REGION Network 5: Procedure Selected
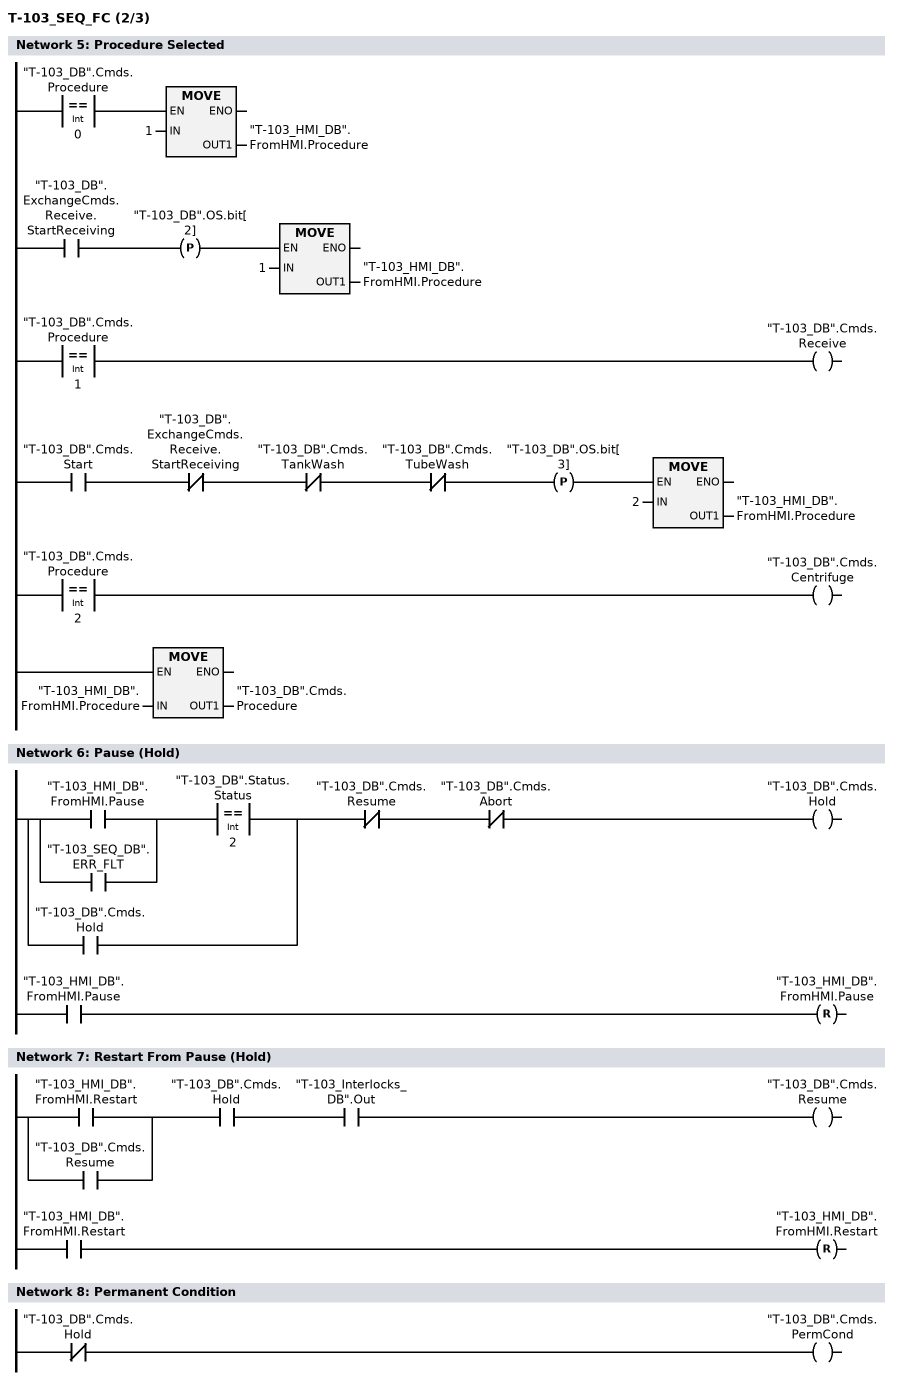
   RUNG wire#powerrail
      { S7_Templates := "SrcType := Int" } EQ_Contact(in1 := "T-103_DB".Cmds.Procedure, in2 := 0)
      Move(in := 1, out1 => "T-103_HMI_DB".FromHMI.Procedure)
   END_RUNG
   RUNG wire#powerrail
      Contact( "T-103_DB".ExchangeCmds.Receive.StartReceiving )
      P_Trig( "T-103_DB".OS.bit[2] )
      Move(in := 1, out1 => "T-103_HMI_DB".FromHMI.Procedure)
   END_RUNG
   RUNG wire#powerrail
      { S7_Templates := "SrcType := Int" } EQ_Contact(in1 := "T-103_DB".Cmds.Procedure, in2 := 1)
      Coil( "T-103_DB".Cmds.Receive )
   END_RUNG
   RUNG wire#powerrail
      Contact( "T-103_DB".Cmds.Start )
      I_Contact( "T-103_DB".ExchangeCmds.Receive.StartReceiving )
      I_Contact( "T-103_DB".Cmds.TankWash )
      I_Contact( "T-103_DB".Cmds.TubeWash )
      P_Trig( "T-103_DB".OS.bit[3] )
      Move(in := 2, out1 => "T-103_HMI_DB".FromHMI.Procedure)
   END_RUNG
   RUNG wire#powerrail
      { S7_Templates := "SrcType := Int" } EQ_Contact(in1 := "T-103_DB".Cmds.Procedure, in2 := 2)
      Coil( "T-103_DB".Cmds.Centrifuge )
   END_RUNG
   RUNG wire#powerrail
      Move(in := "T-103_HMI_DB".FromHMI.Procedure, out1 => "T-103_DB".Cmds.Procedure)
   END_RUNG
   // the same network as SCL:
   IF "T-103_DB".Cmds.Procedure = 0 THEN "T-103_HMI_DB".FromHMI.Procedure := 1; END_IF;
   #_w1 := "T-103_DB".ExchangeCmds.Receive.StartReceiving AND NOT "T-103_DB".OS.bit[2];   // rising edge
   "T-103_DB".OS.bit[2] := "T-103_DB".ExchangeCmds.Receive.StartReceiving;
   IF #_w1 THEN "T-103_HMI_DB".FromHMI.Procedure := 1; END_IF;
   "T-103_DB".Cmds.Receive := "T-103_DB".Cmds.Procedure = 1;
   #_w2 := "T-103_DB".Cmds.Start AND NOT "T-103_DB".ExchangeCmds.Receive.StartReceiving AND NOT "T-103_DB".Cmds.TankWash AND NOT "T-103_DB".Cmds.TubeWash;
   #_w3 := #_w2 AND NOT "T-103_DB".OS.bit[3];   // rising edge
   "T-103_DB".OS.bit[3] := #_w2;
   IF #_w3 THEN "T-103_HMI_DB".FromHMI.Procedure := 2; END_IF;
   "T-103_DB".Cmds.Centrifuge := "T-103_DB".Cmds.Procedure = 2;
   "T-103_DB".Cmds.Procedure := "T-103_HMI_DB".FromHMI.Procedure;
END_REGION

REGION Network 6: Pause (Hold)
   RUNG wire#powerrail
      Contact( "T-103_HMI_DB".FromHMI.Pause )
      wire#w1
      { S7_Templates := "SrcType := Int" } EQ_Contact(in1 := "T-103_DB".Status.Status, in2 := 2)
      wire#w2
      I_Contact( "T-103_DB".Cmds.Resume )
      I_Contact( "T-103_DB".Cmds.Abort )
      Coil( "T-103_DB".Cmds.Hold )
   END_RUNG
   RUNG wire#powerrail
      Contact( "T-103_SEQ_DB".ERR_FLT )
   END_RUNG wire#w1
   RUNG wire#powerrail
      Contact( "T-103_DB".Cmds.Hold )
   END_RUNG wire#w2
   RUNG wire#powerrail
      Contact( "T-103_HMI_DB".FromHMI.Pause )
      R_Coil( "T-103_HMI_DB".FromHMI.Pause )
   END_RUNG
   // the same network as SCL:
   "T-103_DB".Cmds.Hold := ((("T-103_HMI_DB".FromHMI.Pause OR "T-103_SEQ_DB".ERR_FLT) AND ("T-103_DB".Status.Status = 2)) OR "T-103_DB".Cmds.Hold) AND NOT "T-103_DB".Cmds.Resume AND NOT "T-103_DB".Cmds.Abort;
   IF "T-103_HMI_DB".FromHMI.Pause THEN "T-103_HMI_DB".FromHMI.Pause := FALSE; END_IF;
END_REGION

REGION Network 7: Restart From Pause (Hold)
   RUNG wire#powerrail
      Contact( "T-103_HMI_DB".FromHMI.Restart )
      wire#w1
      Contact( "T-103_DB".Cmds.Hold )
      Contact( "T-103_Interlocks_DB".Out )
      Coil( "T-103_DB".Cmds.Resume )
   END_RUNG
   RUNG wire#powerrail
      Contact( "T-103_DB".Cmds.Resume )
   END_RUNG wire#w1
   RUNG wire#powerrail
      Contact( "T-103_HMI_DB".FromHMI.Restart )
      R_Coil( "T-103_HMI_DB".FromHMI.Restart )
   END_RUNG
   // the same network as SCL:
   "T-103_DB".Cmds.Resume := ("T-103_HMI_DB".FromHMI.Restart OR "T-103_DB".Cmds.Resume) AND "T-103_DB".Cmds.Hold AND "T-103_Interlocks_DB".Out;
   IF "T-103_HMI_DB".FromHMI.Restart THEN "T-103_HMI_DB".FromHMI.Restart := FALSE; END_IF;
END_REGION

REGION Network 8: Permanent Condition
   RUNG wire#powerrail
      I_Contact( "T-103_DB".Cmds.Hold )
      Coil( "T-103_DB".Cmds.PermCond )
   END_RUNG
   // the same network as SCL:
   "T-103_DB".Cmds.PermCond := NOT "T-103_DB".Cmds.Hold;
END_REGION

REGION Network 9: Tank Wash
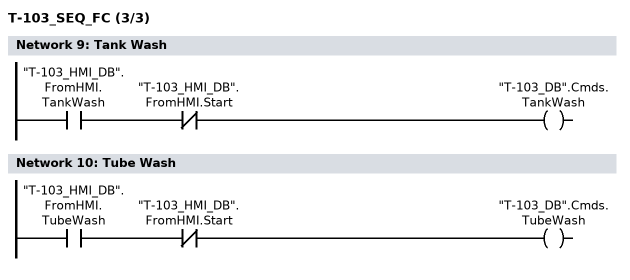
   RUNG wire#powerrail
      Contact( "T-103_HMI_DB".FromHMI.TankWash )
      I_Contact( "T-103_HMI_DB".FromHMI.Start )
      Coil( "T-103_DB".Cmds.TankWash )
   END_RUNG
   // the same network as SCL:
   "T-103_DB".Cmds.TankWash := "T-103_HMI_DB".FromHMI.TankWash AND NOT "T-103_HMI_DB".FromHMI.Start;
END_REGION

REGION Network 10: Tube Wash
   RUNG wire#powerrail
      Contact( "T-103_HMI_DB".FromHMI.TubeWash )
      I_Contact( "T-103_HMI_DB".FromHMI.Start )
      Coil( "T-103_DB".Cmds.TubeWash )
   END_RUNG
   // the same network as SCL:
   "T-103_DB".Cmds.TubeWash := "T-103_HMI_DB".FromHMI.TubeWash AND NOT "T-103_HMI_DB".FromHMI.Start;
END_REGION

REGION Network 11 (SCL): Sequence Status
   IF "T-103_SEQ_DB".S_NO= 1 THEN
       "T-103_DB".Status.Status := 1; //Idle
   ELSIF ("T-103_SEQ_DB".S_NO > 1 AND "T-103_SEQ_DB".S_NO < 150) AND NOT "T-103_SEQ_DB".ERR_FLT AND NOT "T-103_DB".Cmds.Hold THEN
       "T-103_DB".Status.Status := 2; //Running
   ELSIF "T-103_SEQ_DB".S_NO >= 151 AND "T-103_SEQ_DB".S_NO <= 160 AND NOT "T-103_SEQ_DB".ERR_FLT THEN
       "T-103_DB".Status.Status := 3; // Stopping
   ELSIF  "T-103_SEQ_DB".ERR_FLT AND  ("T-103_SEQ_DB".S_NO > 1 AND "T-103_SEQ_DB".S_NO < 150) THEN
       "T-103_DB".Status.Status := 4; // Held
   ELSIF  "T-103_SEQ_DB".ERR_FLT AND  ("T-103_SEQ_DB".S_NO > 1 AND "T-103_SEQ_DB".S_NO < 150) AND "T-103_Aux_DB"."Bool".TOff  THEN
       "T-103_DB".Status.Status := 5; // Holding
   ELSE
       "T-103_DB".Status.Status := 6; // Unknown
   END_IF;

   "T-103_DB".Status.Running := ("T-103_SEQ_DB".S_NO > 3 AND "T-103_SEQ_DB".S_NO <= 150);
   "T-103_DB".Status.Initializing := ("T-103_SEQ_DB".S_NO >= 141 AND "T-103_SEQ_DB".S_NO <= 150);

   //Enable/Disable HMI Start/Stop Button
   "T-103_HMI_DB".ToHMI.EnStopButton := ("T-103_DB".Status.Status > 1) OR "T-103_DB".Status.Step = 0; //Enable HMI Stop Button
   "T-103_HMI_DB".ToHMI.EnStartButton := "T-103_DB".Status.Status = 1; //Idle
   "T-103_HMI_DB".ToHMI.EnPauseButton := "T-103_DB".Status.Status = 2; //Enable Pause Button
   "T-103_HMI_DB".ToHMI.EnRestartButton :=  "T-103_DB".Status.Status = 4; //Enable Restart Button

   //****Interlock Activated
   "T-103_HMI_DB".ToHMI.InterlockActivated := "T-103_Interlocks_DB".Out;
END_REGION

REGION Network 12 (SCL): Sequence Step
   "T-103_DB".Status.Step := "T-103_SEQ_DB".S_NO;
END_REGION

REGION Network 13 (SCL): Sequence state (Procedure running)
   IF "T-103_SEQ_DB".S_NO = 3 OR "T-103_SEQ_DB".S_NO = 4 THEN
       "T-103_DB".Status.State := 1; //Ready
   ELSIF "T-103_SEQ_DB".S_NO >= 21 AND "T-103_SEQ_DB".S_NO <= 60 THEN
       "T-103_DB".Status.State := 2; //Mixing 
   ELSIF "T-103_SEQ_DB".S_NO >= 61 AND "T-103_SEQ_DB".S_NO <= 80 THEN
       "T-103_DB".Status.State := 3; //Pouring
   ELSIF "T-103_SEQ_DB".S_NO >= 141 AND "T-103_SEQ_DB".S_NO <= 150 THEN
       "T-103_DB".Status.State := 4; //Initializing
   ELSIF "T-103_SEQ_DB".S_NO >= 151 AND "T-103_SEQ_DB".S_NO <= 160 THEN
       "T-103_DB".Status.State := 5; //Aborting
   ELSE
       "T-103_DB".Status.State := 0;
   END_IF;
END_REGION

REGION Network 14: Sequence State
END_REGION
END_FUNCTION

// folder: State MACHINE/1)Tanks/Tank T-103 (Cooling Tank)/T-103 <---> Centrifuge

FUNCTION "T-103_Signals_FROM_Centrifuge" : Void   // FC69, LAD
{ S7_Optimized_Access := 'TRUE' }
VERSION : 0.1
BEGIN

REGION Network 1: Start Sequence
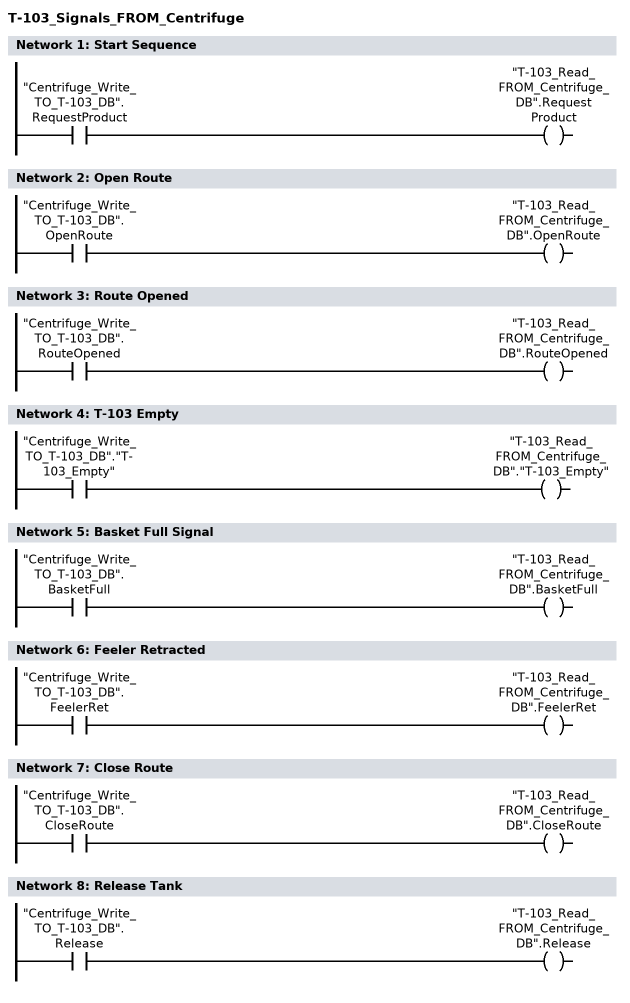
   RUNG wire#powerrail
      Contact( "Centrifuge_Write_TO_T-103_DB".RequestProduct )
      Coil( "T-103_Read_FROM_Centrifuge_DB".RequestProduct )
   END_RUNG
   // the same network as SCL:
   "T-103_Read_FROM_Centrifuge_DB".RequestProduct := "Centrifuge_Write_TO_T-103_DB".RequestProduct;
END_REGION

REGION Network 2: Open Route
   RUNG wire#powerrail
      Contact( "Centrifuge_Write_TO_T-103_DB".OpenRoute )
      Coil( "T-103_Read_FROM_Centrifuge_DB".OpenRoute )
   END_RUNG
   // the same network as SCL:
   "T-103_Read_FROM_Centrifuge_DB".OpenRoute := "Centrifuge_Write_TO_T-103_DB".OpenRoute;
END_REGION

REGION Network 3: Route Opened
   RUNG wire#powerrail
      Contact( "Centrifuge_Write_TO_T-103_DB".RouteOpened )
      Coil( "T-103_Read_FROM_Centrifuge_DB".RouteOpened )
   END_RUNG
   // the same network as SCL:
   "T-103_Read_FROM_Centrifuge_DB".RouteOpened := "Centrifuge_Write_TO_T-103_DB".RouteOpened;
END_REGION

REGION Network 4: T-103 Empty
   RUNG wire#powerrail
      Contact( "Centrifuge_Write_TO_T-103_DB"."T-103_Empty" )
      Coil( "T-103_Read_FROM_Centrifuge_DB"."T-103_Empty" )
   END_RUNG
   // the same network as SCL:
   "T-103_Read_FROM_Centrifuge_DB"."T-103_Empty" := "Centrifuge_Write_TO_T-103_DB"."T-103_Empty";
END_REGION

REGION Network 5: Basket Full Signal
   RUNG wire#powerrail
      Contact( "Centrifuge_Write_TO_T-103_DB".BasketFull )
      Coil( "T-103_Read_FROM_Centrifuge_DB".BasketFull )
   END_RUNG
   // the same network as SCL:
   "T-103_Read_FROM_Centrifuge_DB".BasketFull := "Centrifuge_Write_TO_T-103_DB".BasketFull;
END_REGION

REGION Network 6: Feeler Retracted
   RUNG wire#powerrail
      Contact( "Centrifuge_Write_TO_T-103_DB".FeelerRet )
      Coil( "T-103_Read_FROM_Centrifuge_DB".FeelerRet )
   END_RUNG
   // the same network as SCL:
   "T-103_Read_FROM_Centrifuge_DB".FeelerRet := "Centrifuge_Write_TO_T-103_DB".FeelerRet;
END_REGION

REGION Network 7: Close Route
   RUNG wire#powerrail
      Contact( "Centrifuge_Write_TO_T-103_DB".CloseRoute )
      Coil( "T-103_Read_FROM_Centrifuge_DB".CloseRoute )
   END_RUNG
   // the same network as SCL:
   "T-103_Read_FROM_Centrifuge_DB".CloseRoute := "Centrifuge_Write_TO_T-103_DB".CloseRoute;
END_REGION

REGION Network 8: Release Tank
   RUNG wire#powerrail
      Contact( "Centrifuge_Write_TO_T-103_DB".Release )
      Coil( "T-103_Read_FROM_Centrifuge_DB".Release )
   END_RUNG
   // the same network as SCL:
   "T-103_Read_FROM_Centrifuge_DB".Release := "Centrifuge_Write_TO_T-103_DB".Release;
END_REGION
END_FUNCTION

// folder: State MACHINE/1)Tanks/Tank T-103 (Cooling Tank)/T-103 <---> R-201

FUNCTION "T-103_Signals_FROM_R-201" : Void   // FC49, LAD
{ S7_Optimized_Access := 'TRUE' }
VERSION : 0.1
BEGIN

REGION Network 1: Start Sequence
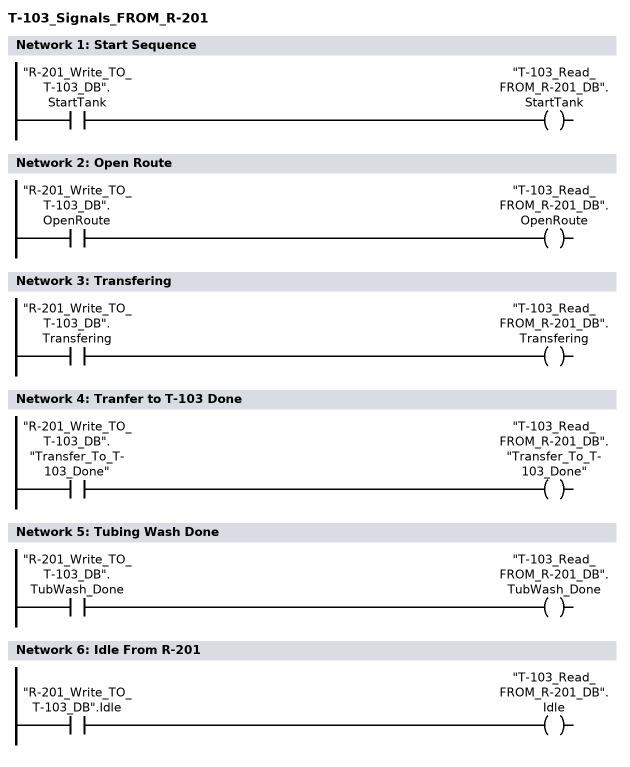
   RUNG wire#powerrail
      Contact( "R-201_Write_TO_T-103_DB".StartTank )
      Coil( "T-103_Read_FROM_R-201_DB".StartTank )
   END_RUNG
   // the same network as SCL:
   "T-103_Read_FROM_R-201_DB".StartTank := "R-201_Write_TO_T-103_DB".StartTank;
END_REGION

REGION Network 2: Open Route
   RUNG wire#powerrail
      Contact( "R-201_Write_TO_T-103_DB".OpenRoute )
      Coil( "T-103_Read_FROM_R-201_DB".OpenRoute )
   END_RUNG
   // the same network as SCL:
   "T-103_Read_FROM_R-201_DB".OpenRoute := "R-201_Write_TO_T-103_DB".OpenRoute;
END_REGION

REGION Network 3: Transfering
   RUNG wire#powerrail
      Contact( "R-201_Write_TO_T-103_DB".Transfering )
      Coil( "T-103_Read_FROM_R-201_DB".Transfering )
   END_RUNG
   // the same network as SCL:
   "T-103_Read_FROM_R-201_DB".Transfering := "R-201_Write_TO_T-103_DB".Transfering;
END_REGION

REGION Network 4: Tranfer to T-103 Done
   RUNG wire#powerrail
      Contact( "R-201_Write_TO_T-103_DB"."Transfer_To_T-103_Done" )
      Coil( "T-103_Read_FROM_R-201_DB"."Transfer_To_T-103_Done" )
   END_RUNG
   // the same network as SCL:
   "T-103_Read_FROM_R-201_DB"."Transfer_To_T-103_Done" := "R-201_Write_TO_T-103_DB"."Transfer_To_T-103_Done";
END_REGION

REGION Network 5: Tubing Wash Done
   RUNG wire#powerrail
      Contact( "R-201_Write_TO_T-103_DB".TubWash_Done )
      Coil( "T-103_Read_FROM_R-201_DB".TubWash_Done )
   END_RUNG
   // the same network as SCL:
   "T-103_Read_FROM_R-201_DB".TubWash_Done := "R-201_Write_TO_T-103_DB".TubWash_Done;
END_REGION

REGION Network 6: Idle From R-201
   RUNG wire#powerrail
      Contact( "R-201_Write_TO_T-103_DB".Idle )
      Coil( "T-103_Read_FROM_R-201_DB".Idle )
   END_RUNG
   // the same network as SCL:
   "T-103_Read_FROM_R-201_DB".Idle := "R-201_Write_TO_T-103_DB".Idle;
END_REGION
END_FUNCTION

// folder: State MACHINE/1)Tanks/Tank T-103 (Cooling Tank)/T-103 <--->R-202

FUNCTION "T-103_Signals_FROM_R-202" : Void   // FC63, LAD
{ S7_Optimized_Access := 'TRUE' }
VERSION : 0.1
BEGIN

REGION Network 1: Start Sequence
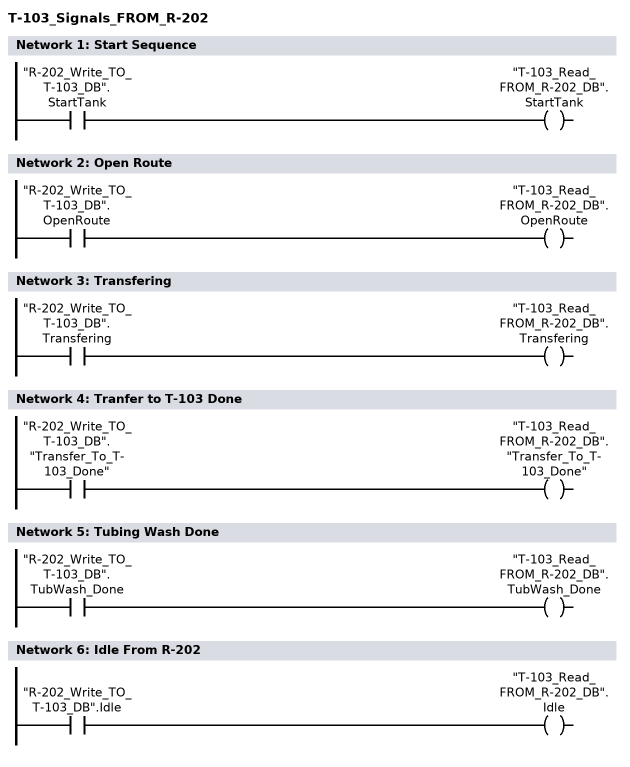
   RUNG wire#powerrail
      Contact( "R-202_Write_TO_T-103_DB".StartTank )
      Coil( "T-103_Read_FROM_R-202_DB".StartTank )
   END_RUNG
   // the same network as SCL:
   "T-103_Read_FROM_R-202_DB".StartTank := "R-202_Write_TO_T-103_DB".StartTank;
END_REGION

REGION Network 2: Open Route
   RUNG wire#powerrail
      Contact( "R-202_Write_TO_T-103_DB".OpenRoute )
      Coil( "T-103_Read_FROM_R-202_DB".OpenRoute )
   END_RUNG
   // the same network as SCL:
   "T-103_Read_FROM_R-202_DB".OpenRoute := "R-202_Write_TO_T-103_DB".OpenRoute;
END_REGION

REGION Network 3: Transfering
   RUNG wire#powerrail
      Contact( "R-202_Write_TO_T-103_DB".Transfering )
      Coil( "T-103_Read_FROM_R-202_DB".Transfering )
   END_RUNG
   // the same network as SCL:
   "T-103_Read_FROM_R-202_DB".Transfering := "R-202_Write_TO_T-103_DB".Transfering;
END_REGION

REGION Network 4: Tranfer to T-103 Done
   RUNG wire#powerrail
      Contact( "R-202_Write_TO_T-103_DB"."Transfer_To_T-103_Done" )
      Coil( "T-103_Read_FROM_R-202_DB"."Transfer_To_T-103_Done" )
   END_RUNG
   // the same network as SCL:
   "T-103_Read_FROM_R-202_DB"."Transfer_To_T-103_Done" := "R-202_Write_TO_T-103_DB"."Transfer_To_T-103_Done";
END_REGION

REGION Network 5: Tubing Wash Done
   RUNG wire#powerrail
      Contact( "R-202_Write_TO_T-103_DB".TubWash_Done )
      Coil( "T-103_Read_FROM_R-202_DB".TubWash_Done )
   END_RUNG
   // the same network as SCL:
   "T-103_Read_FROM_R-202_DB".TubWash_Done := "R-202_Write_TO_T-103_DB".TubWash_Done;
END_REGION

REGION Network 6: Idle From R-202
   RUNG wire#powerrail
      Contact( "R-202_Write_TO_T-103_DB".Idle )
      Coil( "T-103_Read_FROM_R-202_DB".Idle )
   END_RUNG
   // the same network as SCL:
   "T-103_Read_FROM_R-202_DB".Idle := "R-202_Write_TO_T-103_DB".Idle;
END_REGION
END_FUNCTION

// folder: State MACHINE/1)Tanks/Tank T-104 (Water System)

FUNCTION_BLOCK "T-104_SEQ"   // FB38, GRAPH_PLUS
{ S7_Optimized_Access := 'TRUE' }
VERSION : 0.1
   VAR_INPUT
      OFF_SQ : Bool := false;   // Turn sequence off
      INIT_SQ : Bool := false;   // Set sequence to initial state
      ACK_EF : Bool := false;   // Acknowledge all errors and faults
   END_VAR
   VAR_OUTPUT
      S_NO : Int := 0;   // Step number
      S_MORE : Bool := false;   // More steps are available and can be shown in S_NO
      S_ACTIVE : Bool := false;   // Step indicated in S_NO is active
      ERR_FLT : Bool := false;   // Interlock or supervision group error
      AUTO_ON : Bool := false;   // Automatic mode is active
   END_VAR
   VAR
      STATE : Int;   // Current Step in Sequence
      Tank : Struct   // Reactor Ctrl
         IDLE : Bool;
         INITIALIZATION : Bool;   // Sequence initialization
         START : Bool;
         DONE_REACTING : Bool;
         COMPLETE : Bool;   // Reactor Complete Read only
         PARA : Bool;   // PARA load Batch side button
         ABORTING : Bool;   // Sequence about
         WAIT : Bool;   // Wating for Permissive read only
      END_STRUCT;
      TEMP : Struct
         TANKS_BATCH : Real;
         "EMPTY_LV_0%" : Real;
         "MIN_LV_20%" : Real;
         "MAX_LV_80%" : Real;
         "BELOW_32%" : Real;
         "Greater_8%" : Real;
         "PRE-ADD" : Real;
         X_SOL_SIZE : Real;
         Y_SOL_SIZE : Real;
         OFFSEt : Struct
            MAX : Real;
            MIN : Real;
         END_STRUCT;
      END_STRUCT;
      HMI_INFO : Array[0..11] of UInt;
      IF_PAR : G7_IfParPlus_V6;
      RT_DATA : G7_RTDataPlus_V6;   // Internal data area
      Abort : G7_TransitionPlus_V6;   // Transition structure
      InitializeTk : G7_TransitionPlus_V6;   // Transition structure
      Block : G7_TransitionPlus_V6;   // Transition structure
      Rdy : G7_TransitionPlus_V6;   // Transition structure
      Feed : G7_TransitionPlus_V6;   // Transition structure
      ReqWater1 : G7_TransitionPlus_V6;   // Transition structure
      StopWater1 : G7_TransitionPlus_V6;   // Transition structure
      Stoped1 : G7_TransitionPlus_V6;   // Transition structure
      GoBack : G7_TransitionPlus_V6;   // Transition structure
      Init : G7_TransitionPlus_V6;   // Transition structure
      SAut : G7_TransitionPlus_V6;   // Transition structure
      SIn : G7_TransitionPlus_V6;   // Transition structure
      Initd : G7_TransitionPlus_V6;   // Transition structure
      Ab : G7_TransitionPlus_V6;   // Transition structure
      AbortOn : G7_TransitionPlus_V6;   // Transition structure
      DneAbort : G7_TransitionPlus_V6;   // Transition structure
      Idle : G7_StepPlus_V6;   // Step structure
      Ready : G7_StepPlus_V6;   // Step structure
      SelectSeq : G7_StepPlus_V6;   // Step structure
      FeedStarted : G7_StepPlus_V6;   // Step structure
      Feeding : G7_StepPlus_V6;   // Step structure
      StopTransfer : G7_StepPlus_V6;   // Step structure
      Done : G7_StepPlus_V6;   // Step structure
      Initialize : G7_StepPlus_V6;   // Step structure
      SetAuto : G7_StepPlus_V6;   // Step structure
      SetInitial : G7_StepPlus_V6;   // Step structure
      Initialized : G7_StepPlus_V6;   // Step structure
      AbortStarting : G7_StepPlus_V6;   // Step structure
      Aborting : G7_StepPlus_V6;   // Step structure
      Abort_Done : G7_StepPlus_V6;   // Step structure
      SINI : Array[0..4] of USInt;
      LSTT : Array[0..15] of USInt;
      ATAJ : Array[0..15] of USInt;
      ATAB : Array[0..15] of USInt;
      PSTT : Array[0..15] of USInt;
      NSTT : Array[0..15] of USInt;
      ASSJ : Array[0..13] of USInt;
      ASSB : Array[0..13] of USInt;
      PTTS : Array[0..13] of USInt;
      NTTS : Array[0..13] of USInt;
      SW_SQTS : Array[0..13] of USInt;
      SWITCH : Array[0..3] of USInt;
      TVX : Array[0..7] of USInt;
      TTX : Array[0..7] of USInt;
      TSX : Array[0..4] of USInt;
      S00X : Array[0..4] of USInt;
      SOFFX : Array[0..4] of USInt;
      SONX : Array[0..4] of USInt;
      SAX : Array[0..4] of USInt;
      SERRX : Array[0..14] of USInt;
      SMX : Array[0..14] of USInt;
      S0X : Array[0..14] of USInt;
      S1X : Array[0..14] of USInt;
      IL_ALARM_INST : Diag_Alarm;
      SUP_ALARM_INST : Diag_Alarm;
      STEP_TIME_ALARM_INST : Diag_Alarm;
      IEC_TIMER_INST : IEC_TIMER;
      TRANSACTION_FLAG : Bool := false;
   END_VAR
   VAR CONSTANT
      "Single R-201 T-101 seq done" : Int := 214;
      "Single R-201 T-102 seq done" : Int := 218;
   END_VAR
   // SINI[0] := 2;
   // LSTT[0] := 11;
   // NSTT[0] := 11;
   // PTTS[0] := 255;
   // TVX[0] := 16#1;
   // TTX[0] := 16#1;
   // TSX[0] := 16#1;
   // S00X[0] := 16#1;
   // SOFFX[0] := 16#1;
   // SONX[0] := 16#1;
   // SAX[0] := 16#1;
   // SERRX[0] := 16#1;
   // SMX[0] := 16#1;
   // S0X[0] := 16#1;
   // S1X[0] := 16#1;
   // LSTT[1] := 7;
   // LSTT[2] := 255;
   // LSTT[3] := 255;
   // LSTT[4] := 3;
   // LSTT[5] := 255;
   // LSTT[6] := 255;
   // LSTT[7] := 255;
   // LSTT[8] := 3;
   // LSTT[9] := 255;
   // LSTT[10] := 255;
   // LSTT[11] := 255;
   // LSTT[13] := 255;
   // ATAJ[1] := 1;
   // ATAJ[2] := 2;
   // ATAJ[3] := 3;
   // ATAJ[4] := 4;
   // ATAJ[5] := 5;
   // ATAJ[6] := 6;
   // ATAJ[7] := 7;
   // ATAJ[8] := 8;
   // ATAJ[9] := 9;
   // ATAJ[10] := 10;
   // ATAJ[11] := 11;
   // ATAJ[12] := 12;
   // ATAJ[13] := 13;
   // ATAB[1] := 2;
   // ATAB[13] := 13;
   // ATAB[3] := 3;
   // ATAB[4] := 4;
   // ATAB[5] := 5;
   // ATAB[6] := 6;
   // ATAB[7] := 7;
   // ATAB[8] := 8;
   // ATAB[9] := 9;
   // ATAB[10] := 10;
   // ATAB[11] := 11;
   // ATAB[12] := 12;
   // PSTT[3] := 1;
   // PSTT[4] := 2;
   // PSTT[5] := 3;
   // PSTT[6] := 4;
   // PSTT[7] := 5;
   // PSTT[8] := 6;
   // PSTT[9] := 7;
   // PSTT[10] := 8;
   // PSTT[11] := 9;
   // PSTT[12] := 10;
   // NSTT[1] := 7;
   // NSTT[2] := 1;
   // NSTT[3] := 2;
   // NSTT[4] := 3;
   // NSTT[5] := 4;
   // NSTT[6] := 5;
   // NSTT[7] := 6;
   // NSTT[8] := 3;
   // NSTT[9] := 8;
   // NSTT[10] := 9;
   // NSTT[11] := 10;
   // NSTT[13] := 12;
   // ASSJ[1] := 1;
   // ASSJ[2] := 2;
   // ASSJ[3] := 3;
   // ASSJ[4] := 4;
   // ASSJ[5] := 5;
   // ASSJ[6] := 6;
   // ASSJ[7] := 7;
   // ASSJ[8] := 8;
   // ASSJ[9] := 9;
   // ASSJ[10] := 10;
   // ASSJ[11] := 11;
   // ASSB[1] := 1;
   // ASSB[2] := 2;
   // ASSB[3] := 3;
   // ASSB[4] := 4;
   // ASSB[5] := 5;
   // ASSB[6] := 6;
   // ASSB[7] := 7;
   // ASSB[8] := 8;
   // ASSB[9] := 9;
   // ASSB[10] := 10;
   // ASSB[11] := 11;
   // PTTS[4] := 5;
   // PTTS[3] := 255;
   // PTTS[5] := 6;
   // PTTS[6] := 7;
   // PTTS[7] := 255;
   // PTTS[8] := 9;
   // PTTS[9] := 10;
   // PTTS[11] := 255;
   // SW_SQTS[4] := 2;
   // NTTS[2] := 4;
   // NTTS[3] := 5;
   // NTTS[4] := 6;
   // NTTS[5] := 7;
   // NTTS[6] := 8;
   // NTTS[7] := 9;
   // NTTS[8] := 10;
   // NTTS[9] := 11;
   // NTTS[10] := 12;
   // NTTS[11] := 13;
   // SW_SQTS[5] := 2;
   // SW_SQTS[8] := 3;
   // SW_SQTS[9] := 3;
   // SW_SQTS[11] := 4;
   // SWITCH[0] := 156;
   // SWITCH[2] := 251;
   // PSTT[13] := 11;
   // PTTS[1] := 2;
   // NTTS[1] := 3;
   // SW_SQTS[1] := 1;
   // PTTS[10] := 11;
   // ATAB[0] := 1;
   // SINI[4] := 255;
   // SINI[3] := 255;
   // PTTS[2] := 3;
   // SW_SQTS[7] := 3;
   // SW_SQTS[6] := 2;
   // SWITCH[1] := 239;
   // SINI[2] := 255;
   // SW_SQTS[3] := 2;
   // SW_SQTS[2] := 1;
   // SW_SQTS[10] := 3;
   // LSTT[12] := 1;
   // LSTT[14] := 255;
   // ATAJ[14] := 14;
   // ATAJ[15] := 15;
   // ATAB[14] := 14;
   // ATAB[15] := 15;
   // PSTT[14] := 12;
   // PSTT[15] := 13;
   // NSTT[12] := 1;
   // NSTT[14] := 13;
   // ASSJ[12] := 12;
   // ASSJ[13] := 13;
   // ASSB[12] := 12;
   // ASSB[13] := 13;
   // PTTS[12] := 13;
   // PTTS[13] := 14;
   // NTTS[12] := 14;
   // NTTS[13] := 15;
   // SW_SQTS[12] := 4;
   // SW_SQTS[13] := 4;
BEGIN
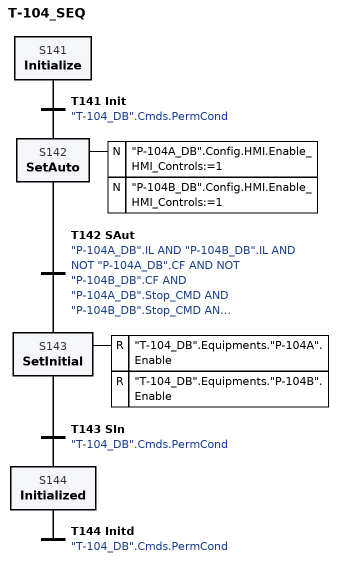
   // permanent pre-instructions
   NETWORK 1
      "T-104_SEQ_FC"();
      "T-104_Signals_FROM_R-201"();
      "T-104_Signals_FROM_R-202"();
      "T-104_Signals_FROM_T-101"();
      "T-104_Signals_FROM_T-102"();
      "T-104_Signals_FROM_Centrifuge"();
      "T-104_SignalsInExchange"();

   // sequencer 1
   STEP SetAuto:   // S142, max time T#10S, warning time T#7S
      // PMP OFF
              N    "P-104A_DB".Config.HMI.Enable_HMI_Controls:=1
              N    "P-104B_DB".Config.HMI.Enable_HMI_Controls:=1
   END_STEP
   TRANSITION SAut FROM SetAuto TO SetInitial   // T142: OFF: P-101A/B
      := "P-104A_DB".IL AND "P-104B_DB".IL AND NOT "P-104A_DB".CF AND NOT "P-104B_DB".CF AND "P-104A_DB".Stop_CMD AND "P-104B_DB".Stop_CMD AND "T-104_DB".Cmds.PermCond;
   END_TRANSITION
   STEP Initialize:   // S141, max time T#10S, warning time T#7S
   END_STEP
   TRANSITION Init FROM Initialize TO SetAuto   // T141
      := "T-104_DB".Cmds.PermCond;
   END_TRANSITION
   STEP SetInitial:   // S143, max time T#10S, warning time T#7S
              R    "T-104_DB".Equipments."P-104A".Enable
              R    "T-104_DB".Equipments."P-104B".Enable
   END_STEP
   TRANSITION SIn FROM SetInitial TO Initialized   // T143
      := "T-104_DB".Cmds.PermCond;
   END_TRANSITION
   STEP Initialized:   // S144, max time T#10S, warning time T#7S
   END_STEP
   TRANSITION Initd FROM Initialized TO ?   // T144
      := "T-104_DB".Cmds.PermCond;
   END_TRANSITION

   // permanent post-instructions
   NETWORK 1
      "T-104_SignalsOutExchange"();
      "T-104_FC_Outputs"();
END_FUNCTION_BLOCK

FUNCTION "T-104_SignalsInExchange" : Void   // FC52, LAD
{ S7_Optimized_Access := 'TRUE' }
VERSION : 0.1
BEGIN

REGION Network 1: Start (Receive)
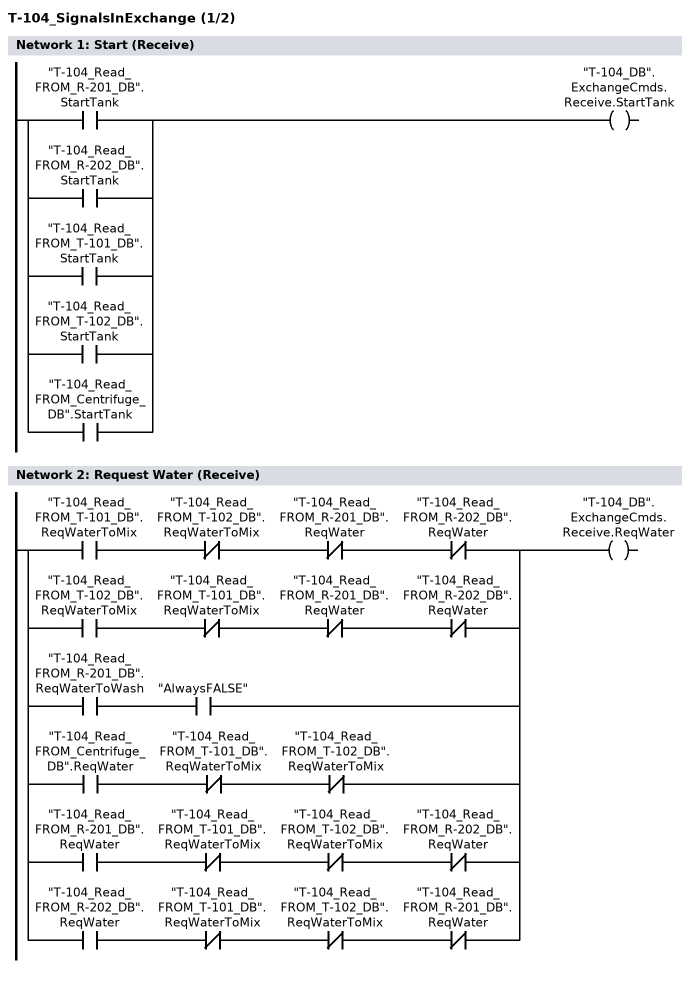
   RUNG wire#powerrail
      Contact( "T-104_Read_FROM_R-201_DB".StartTank )
      wire#w1
      Coil( "T-104_DB".ExchangeCmds.Receive.StartTank )
   END_RUNG
   RUNG wire#powerrail
      Contact( "T-104_Read_FROM_R-202_DB".StartTank )
   END_RUNG wire#w1
   RUNG wire#powerrail
      Contact( "T-104_Read_FROM_T-101_DB".StartTank )
   END_RUNG wire#w1
   RUNG wire#powerrail
      Contact( "T-104_Read_FROM_T-102_DB".StartTank )
   END_RUNG wire#w1
   RUNG wire#powerrail
      Contact( "T-104_Read_FROM_Centrifuge_DB".StartTank )
   END_RUNG wire#w1
   // the same network as SCL:
   "T-104_DB".ExchangeCmds.Receive.StartTank := "T-104_Read_FROM_R-201_DB".StartTank OR "T-104_Read_FROM_R-202_DB".StartTank OR "T-104_Read_FROM_T-101_DB".StartTank OR "T-104_Read_FROM_T-102_DB".StartTank OR "T-104_Read_FROM_Centrifuge_DB".StartTank;
END_REGION

REGION Network 2: Request Water (Receive)
   RUNG wire#powerrail
      Contact( "T-104_Read_FROM_T-101_DB".ReqWaterToMix )
      I_Contact( "T-104_Read_FROM_T-102_DB".ReqWaterToMix )
      I_Contact( "T-104_Read_FROM_R-201_DB".ReqWater )
      I_Contact( "T-104_Read_FROM_R-202_DB".ReqWater )
      wire#w1
      Coil( "T-104_DB".ExchangeCmds.Receive.ReqWater )
   END_RUNG
   RUNG wire#powerrail
      Contact( "T-104_Read_FROM_T-102_DB".ReqWaterToMix )
      I_Contact( "T-104_Read_FROM_T-101_DB".ReqWaterToMix )
      I_Contact( "T-104_Read_FROM_R-201_DB".ReqWater )
      I_Contact( "T-104_Read_FROM_R-202_DB".ReqWater )
   END_RUNG wire#w1
   RUNG wire#powerrail
      Contact( "T-104_Read_FROM_R-201_DB".ReqWaterToWash )
      Contact( "AlwaysFALSE" )
   END_RUNG wire#w1
   RUNG wire#powerrail
      Contact( "T-104_Read_FROM_Centrifuge_DB".ReqWater )
      I_Contact( "T-104_Read_FROM_T-101_DB".ReqWaterToMix )
      I_Contact( "T-104_Read_FROM_T-102_DB".ReqWaterToMix )
   END_RUNG wire#w1
   RUNG wire#powerrail
      Contact( "T-104_Read_FROM_R-201_DB".ReqWater )
      I_Contact( "T-104_Read_FROM_T-101_DB".ReqWaterToMix )
      I_Contact( "T-104_Read_FROM_T-102_DB".ReqWaterToMix )
      I_Contact( "T-104_Read_FROM_R-202_DB".ReqWater )
   END_RUNG wire#w1
   RUNG wire#powerrail
      Contact( "T-104_Read_FROM_R-202_DB".ReqWater )
      I_Contact( "T-104_Read_FROM_T-101_DB".ReqWaterToMix )
      I_Contact( "T-104_Read_FROM_T-102_DB".ReqWaterToMix )
      I_Contact( "T-104_Read_FROM_R-201_DB".ReqWater )
   END_RUNG wire#w1
   // the same network as SCL:
   "T-104_DB".ExchangeCmds.Receive.ReqWater := ("T-104_Read_FROM_T-101_DB".ReqWaterToMix AND NOT "T-104_Read_FROM_T-102_DB".ReqWaterToMix AND NOT "T-104_Read_FROM_R-201_DB".ReqWater AND NOT "T-104_Read_FROM_R-202_DB".ReqWater) OR ("T-104_Read_FROM_T-102_DB".ReqWaterToMix AND NOT "T-104_Read_FROM_T-101_DB".ReqWaterToMix AND NOT "T-104_Read_FROM_R-201_DB".ReqWater AND NOT "T-104_Read_FROM_R-202_DB".ReqWater) OR ("T-104_Read_FROM_R-201_DB".ReqWaterToWash AND "AlwaysFALSE") OR ("T-104_Read_FROM_Centrifuge_DB".ReqWater AND NOT "T-104_Read_FROM_T-101_DB".ReqWaterToMix AND NOT "T-104_Read_FROM_T-102_DB".ReqWaterToMix) OR ("T-104_Read_FROM_R-201_DB".ReqWater AND NOT "T-104_Read_FROM_T-101_DB".ReqWaterToMix AND NOT "T-104_Read_FROM_T-102_DB".ReqWaterToMix AND NOT "T-104_Read_FROM_R-202_DB".ReqWater) OR ("T-104_Read_FROM_R-202_DB".ReqWater AND NOT "T-104_Read_FROM_T-101_DB".ReqWaterToMix AND NOT "T-104_Read_FROM_T-102_DB".ReqWaterToMix AND NOT "T-104_Read_FROM_R-201_DB".ReqWater);
END_REGION

REGION Network 3: Stop Request Water (Receive)
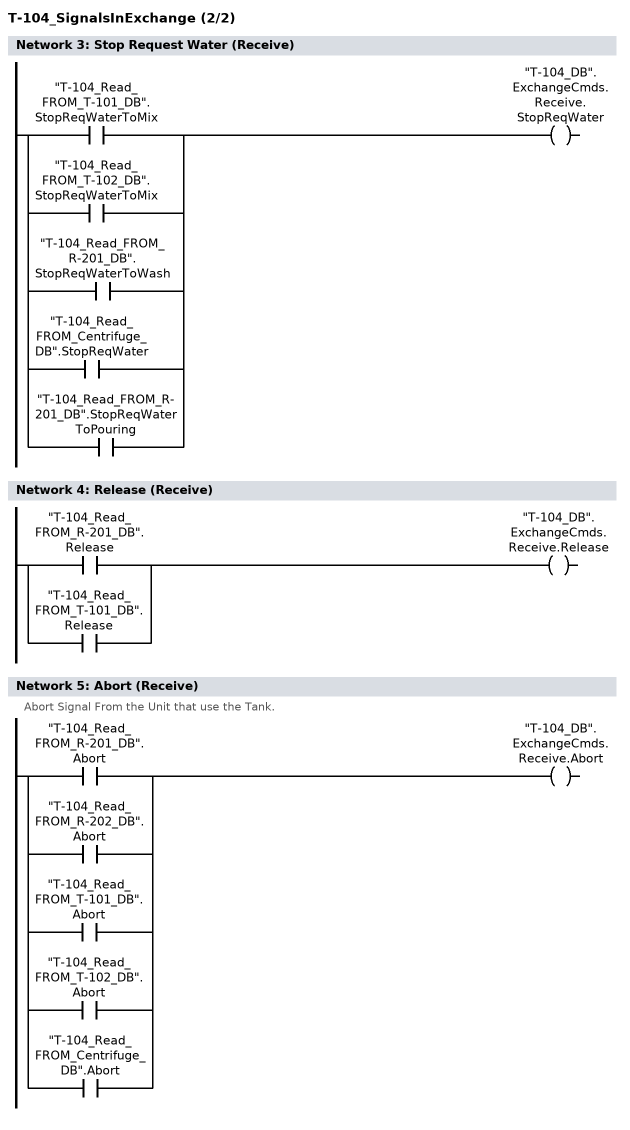
   RUNG wire#powerrail
      Contact( "T-104_Read_FROM_T-101_DB".StopReqWaterToMix )
      wire#w1
      Coil( "T-104_DB".ExchangeCmds.Receive.StopReqWater )
   END_RUNG
   RUNG wire#powerrail
      Contact( "T-104_Read_FROM_T-102_DB".StopReqWaterToMix )
   END_RUNG wire#w1
   RUNG wire#powerrail
      Contact( "T-104_Read_FROM_R-201_DB".StopReqWaterToWash )
   END_RUNG wire#w1
   RUNG wire#powerrail
      Contact( "T-104_Read_FROM_Centrifuge_DB".StopReqWater )
   END_RUNG wire#w1
   RUNG wire#powerrail
      Contact( "T-104_Read_FROM_R-201_DB".StopReqWaterToPouring )
   END_RUNG wire#w1
   // the same network as SCL:
   "T-104_DB".ExchangeCmds.Receive.StopReqWater := "T-104_Read_FROM_T-101_DB".StopReqWaterToMix OR "T-104_Read_FROM_T-102_DB".StopReqWaterToMix OR "T-104_Read_FROM_R-201_DB".StopReqWaterToWash OR "T-104_Read_FROM_Centrifuge_DB".StopReqWater OR "T-104_Read_FROM_R-201_DB".StopReqWaterToPouring;
END_REGION

REGION Network 4: Release (Receive)
   RUNG wire#powerrail
      Contact( "T-104_Read_FROM_R-201_DB".Release )
      wire#w1
      Coil( "T-104_DB".ExchangeCmds.Receive.Release )
   END_RUNG
   RUNG wire#powerrail
      Contact( "T-104_Read_FROM_T-101_DB".Release )
   END_RUNG wire#w1
   // the same network as SCL:
   "T-104_DB".ExchangeCmds.Receive.Release := "T-104_Read_FROM_R-201_DB".Release OR "T-104_Read_FROM_T-101_DB".Release;
END_REGION

REGION Network 5: Abort (Receive)
   // Abort Signal From the Unit that use the Tank.
   RUNG wire#powerrail
      Contact( "T-104_Read_FROM_R-201_DB".Abort )
      wire#w1
      Coil( "T-104_DB".ExchangeCmds.Receive.Abort )
   END_RUNG
   RUNG wire#powerrail
      Contact( "T-104_Read_FROM_R-202_DB".Abort )
   END_RUNG wire#w1
   RUNG wire#powerrail
      Contact( "T-104_Read_FROM_T-101_DB".Abort )
   END_RUNG wire#w1
   RUNG wire#powerrail
      Contact( "T-104_Read_FROM_T-102_DB".Abort )
   END_RUNG wire#w1
   RUNG wire#powerrail
      Contact( "T-104_Read_FROM_Centrifuge_DB".Abort )
   END_RUNG wire#w1
   // the same network as SCL:
   "T-104_DB".ExchangeCmds.Receive.Abort := "T-104_Read_FROM_R-201_DB".Abort OR "T-104_Read_FROM_R-202_DB".Abort OR "T-104_Read_FROM_T-101_DB".Abort OR "T-104_Read_FROM_T-102_DB".Abort OR "T-104_Read_FROM_Centrifuge_DB".Abort;
END_REGION
END_FUNCTION

FUNCTION "T-104_FC_Outputs" : Void   // FC79, SCL
{ S7_Optimized_Access := 'TRUE' }